(* Logix 5000 project; controller PLC_MCC1300_75F1 vendor 1 type 14 code 166 rev 32.11; software revision 32.04; part 41 of 83 *)
(* tags used below, declared in another part *)
   GP_RampSpace : GP_RampSpace;
   I : INT[128];   // Local Input Updates Input Slot 2
   TMP_d : DINT;
   TMP_dConv : DINT;
   TMP_dConvDebug : DINT;
   TMP_dEndConveyorPos : DINT;
   TMP_dIndexNext : DINT;
   TMP_dIndexNextDebug : DINT;
   TMP_dIndexPreviousDebug : DINT;
   TMP_dTailOnNextConveyor_cmm : DINT;
   TMP_xLastConvDebug : BOOL;
   TMP_xOSN : DINT;
   TMP_xOSN_B : DINT;
   TMP_xOSR : DINT;
   TMP_xOSR_B : DINT;
   xAlwaysOFF : BOOL;
   xAlwaysON : BOOL;
   xDebugOFF : BOOL;
   xDebugON : BOOL;
   Z300_Conveyor : UDT_StandConv[29];
   Z300_Conveyor_ALM : MAC_Conveyor_ZC_ALM[29];
   Z300_Conveyor_Conf : UDT_Conveyor_Config[29];
   Z300_Conveyor_HMR : MAC_Conveyor_ZC_HMR[29];
   Z300_Conveyor_HMW : MAC_Conveyor_ZC_HMW[29];
   Z300_LineTracking : UDT_LINE_TRACKING;
(* MainProgram, continued *)

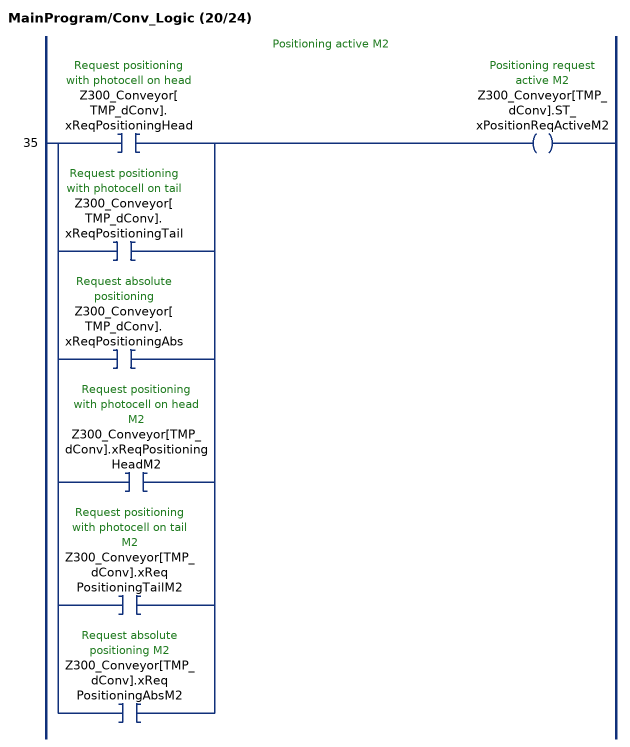
   // Positioning active M2
   35: [XIC(Z300_Conveyor[TMP_dConv].xReqPositioningHead) ,XIC(Z300_Conveyor[TMP_dConv].xReqPositioningTail) ,XIC(Z300_Conveyor[TMP_dConv].xReqPositioningAbs) ,XIC(Z300_Conveyor[TMP_dConv].xReqPositioningHeadM2) ,XIC(Z300_Conveyor[TMP_dConv].xReqPositioningTailM2) ,XIC(Z300_Conveyor[TMP_dConv].xReqPositioningAbsM2) ]OTE(Z300_Conveyor[TMP_dConv].ST_xPositionReqActiveM2);
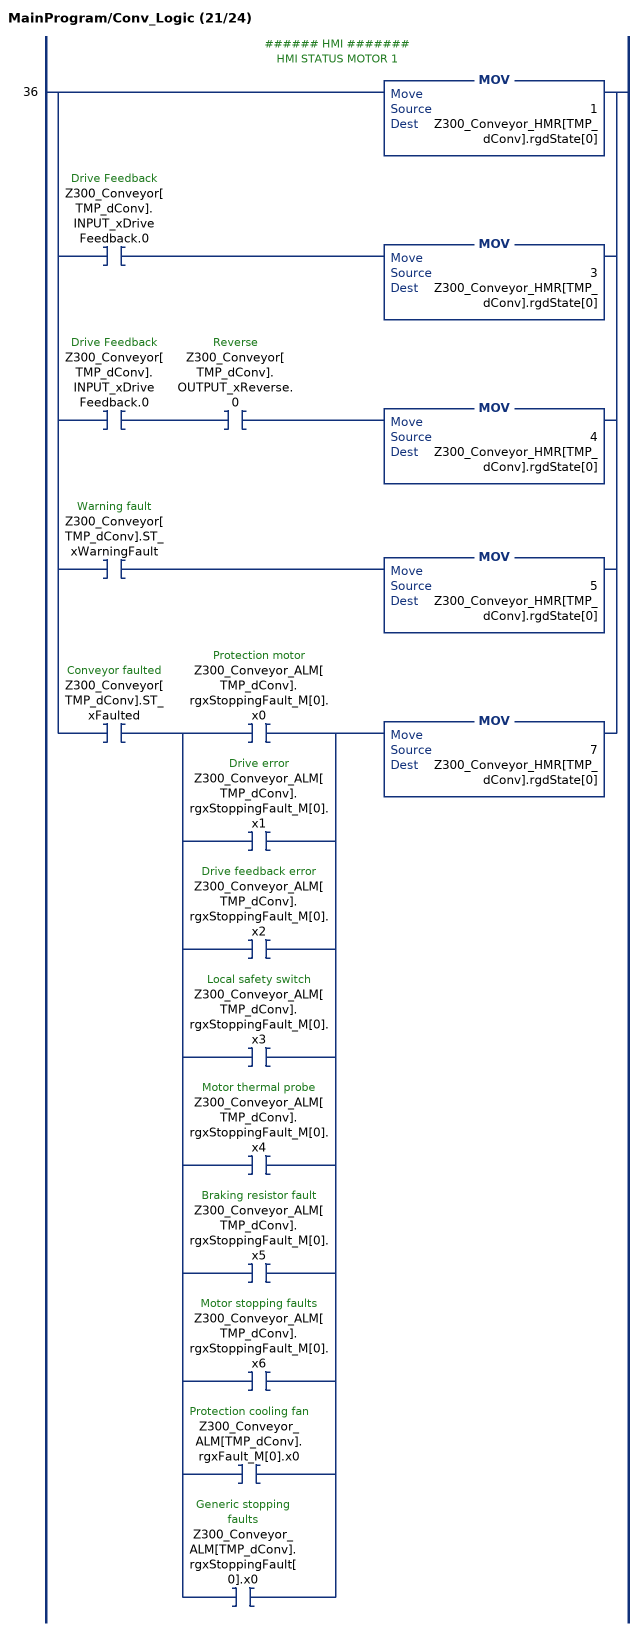
   // ###### HMI #######
   // HMI STATUS MOTOR 1
   36: [MOV(1,Z300_Conveyor_HMR[TMP_dConv].rgdState[0]) ,XIC(Z300_Conveyor[TMP_dConv].INPUT_xDriveFeedback.0) MOV(3,Z300_Conveyor_HMR[TMP_dConv].rgdState[0]) ,XIC(Z300_Conveyor[TMP_dConv].INPUT_xDriveFeedback.0) XIC(Z300_Conveyor[TMP_dConv].OUTPUT_xReverse.0) MOV(4,Z300_Conveyor_HMR[TMP_dConv].rgdState[0]) ,XIC(Z300_Conveyor[TMP_dConv].ST_xWarningFault) MOV(5,Z300_Conveyor_HMR[TMP_dConv].rgdState[0]) ,XIC(Z300_Conveyor[TMP_dConv].ST_xFaulted) [XIC(Z300_Conveyor_ALM[TMP_dConv].rgxStoppingFault_M[0].x0) ,XIC(Z300_Conveyor_ALM[TMP_dConv].rgxStoppingFault_M[0].x1) ,XIC(Z300_Conveyor_ALM[TMP_dConv].rgxStoppingFault_M[0].x2) ,XIC(Z300_Conveyor_ALM[TMP_dConv].rgxStoppingFault_M[0].x3) ,XIC(Z300_Conveyor_ALM[TMP_dConv].rgxStoppingFault_M[0].x4) ,XIC(Z300_Conveyor_ALM[TMP_dConv].rgxStoppingFault_M[0].x5) ,XIC(Z300_Conveyor_ALM[TMP_dConv].rgxStoppingFault_M[0].x6) ,XIC(Z300_Conveyor_ALM[TMP_dConv].rgxFault_M[0].x0) ,XIC(Z300_Conveyor_ALM[TMP_dConv].rgxStoppingFault[0].x0) ] MOV(7,Z300_Conveyor_HMR[TMP_dConv].rgdState[0]) ];
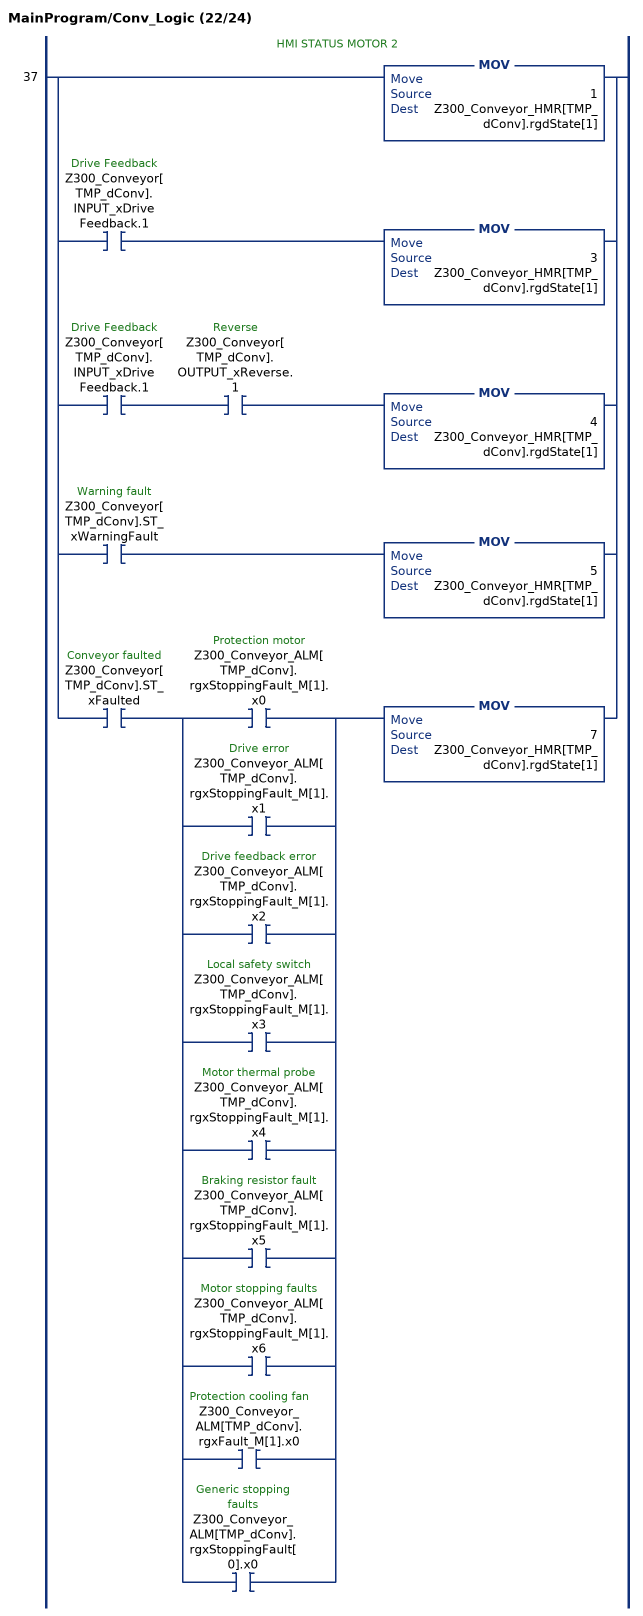
   // HMI STATUS MOTOR 2
   37: [MOV(1,Z300_Conveyor_HMR[TMP_dConv].rgdState[1]) ,XIC(Z300_Conveyor[TMP_dConv].INPUT_xDriveFeedback.1) MOV(3,Z300_Conveyor_HMR[TMP_dConv].rgdState[1]) ,XIC(Z300_Conveyor[TMP_dConv].INPUT_xDriveFeedback.1) XIC(Z300_Conveyor[TMP_dConv].OUTPUT_xReverse.1) MOV(4,Z300_Conveyor_HMR[TMP_dConv].rgdState[1]) ,XIC(Z300_Conveyor[TMP_dConv].ST_xWarningFault) MOV(5,Z300_Conveyor_HMR[TMP_dConv].rgdState[1]) ,XIC(Z300_Conveyor[TMP_dConv].ST_xFaulted) [XIC(Z300_Conveyor_ALM[TMP_dConv].rgxStoppingFault_M[1].x0) ,XIC(Z300_Conveyor_ALM[TMP_dConv].rgxStoppingFault_M[1].x1) ,XIC(Z300_Conveyor_ALM[TMP_dConv].rgxStoppingFault_M[1].x2) ,XIC(Z300_Conveyor_ALM[TMP_dConv].rgxStoppingFault_M[1].x3) ,XIC(Z300_Conveyor_ALM[TMP_dConv].rgxStoppingFault_M[1].x4) ,XIC(Z300_Conveyor_ALM[TMP_dConv].rgxStoppingFault_M[1].x5) ,XIC(Z300_Conveyor_ALM[TMP_dConv].rgxStoppingFault_M[1].x6) ,XIC(Z300_Conveyor_ALM[TMP_dConv].rgxFault_M[1].x0) ,XIC(Z300_Conveyor_ALM[TMP_dConv].rgxStoppingFault[0].x0) ] MOV(7,Z300_Conveyor_HMR[TMP_dConv].rgdState[1]) ];
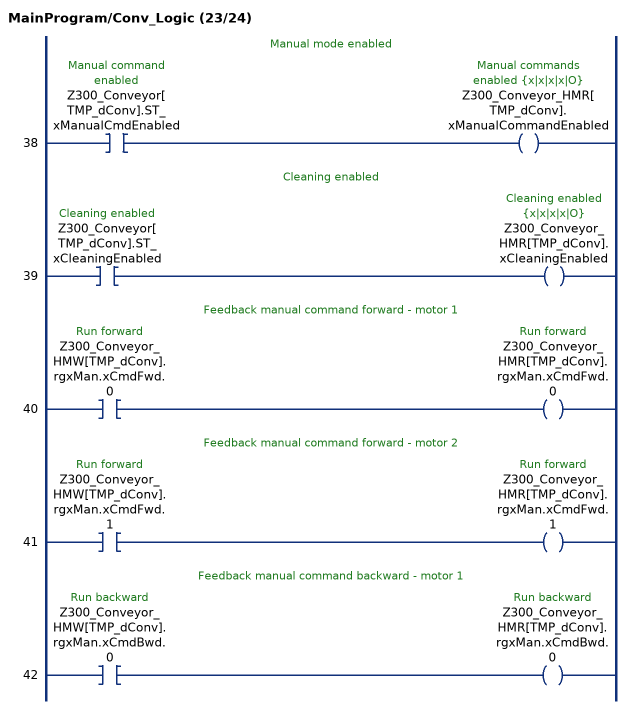
   // Manual mode enabled
   38: XIC(Z300_Conveyor[TMP_dConv].ST_xManualCmdEnabled)OTE(Z300_Conveyor_HMR[TMP_dConv].xManualCommandEnabled);
   // Cleaning enabled
   39: XIC(Z300_Conveyor[TMP_dConv].ST_xCleaningEnabled)OTE(Z300_Conveyor_HMR[TMP_dConv].xCleaningEnabled);
   // Feedback manual command forward - motor 1
   40: XIC(Z300_Conveyor_HMW[TMP_dConv].rgxMan.xCmdFwd.0)OTE(Z300_Conveyor_HMR[TMP_dConv].rgxMan.xCmdFwd.0);
   // Feedback manual command forward - motor 2
   41: XIC(Z300_Conveyor_HMW[TMP_dConv].rgxMan.xCmdFwd.1)OTE(Z300_Conveyor_HMR[TMP_dConv].rgxMan.xCmdFwd.1);
   // Feedback manual command backward - motor 1
   42: XIC(Z300_Conveyor_HMW[TMP_dConv].rgxMan.xCmdBwd.0)OTE(Z300_Conveyor_HMR[TMP_dConv].rgxMan.xCmdBwd.0);
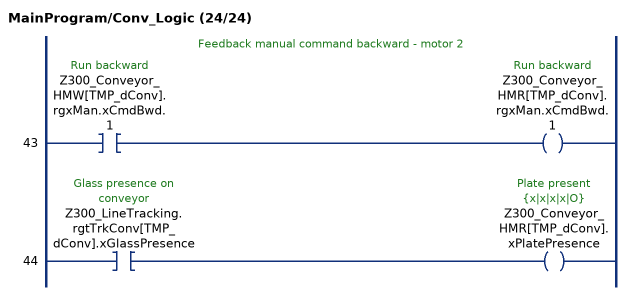
   // Feedback manual command backward - motor 2
   43: XIC(Z300_Conveyor_HMW[TMP_dConv].rgxMan.xCmdBwd.1)OTE(Z300_Conveyor_HMR[TMP_dConv].rgxMan.xCmdBwd.1);
   44: XIC(Z300_LineTracking.rgtTrkConv[TMP_dConv].xGlassPresence)OTE(Z300_Conveyor_HMR[TMP_dConv].xPlatePresence);
END_ROUTINE

ROUTINE Conv_Logic_Debug   (* ladder *)
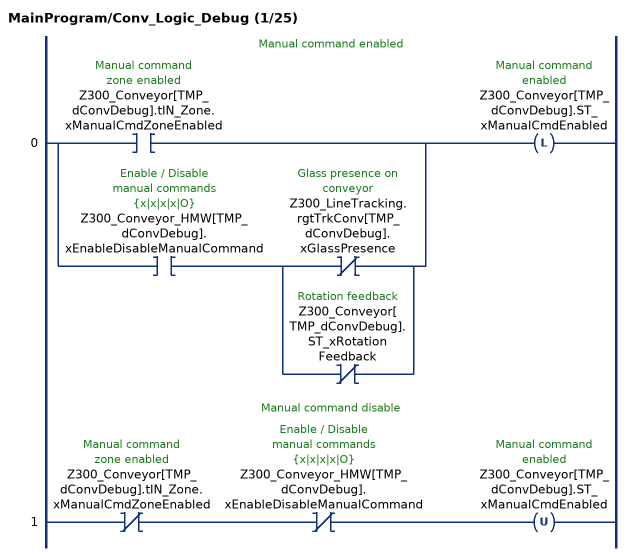
   // Manual command enabled
   0: [XIC(Z300_Conveyor[TMP_dConvDebug].tIN_Zone.xManualCmdZoneEnabled) ,XIC(Z300_Conveyor_HMW[TMP_dConvDebug].xEnableDisableManualCommand) [XIO(Z300_LineTracking.rgtTrkConv[TMP_dConvDebug].xGlassPresence) ,XIO(Z300_Conveyor[TMP_dConvDebug].ST_xRotationFeedback) ] ]OTL(Z300_Conveyor[TMP_dConvDebug].ST_xManualCmdEnabled);
   // Manual command disable
   1: XIO(Z300_Conveyor[TMP_dConvDebug].tIN_Zone.xManualCmdZoneEnabled)XIO(Z300_Conveyor_HMW[TMP_dConvDebug].xEnableDisableManualCommand)OTU(Z300_Conveyor[TMP_dConvDebug].ST_xManualCmdEnabled);
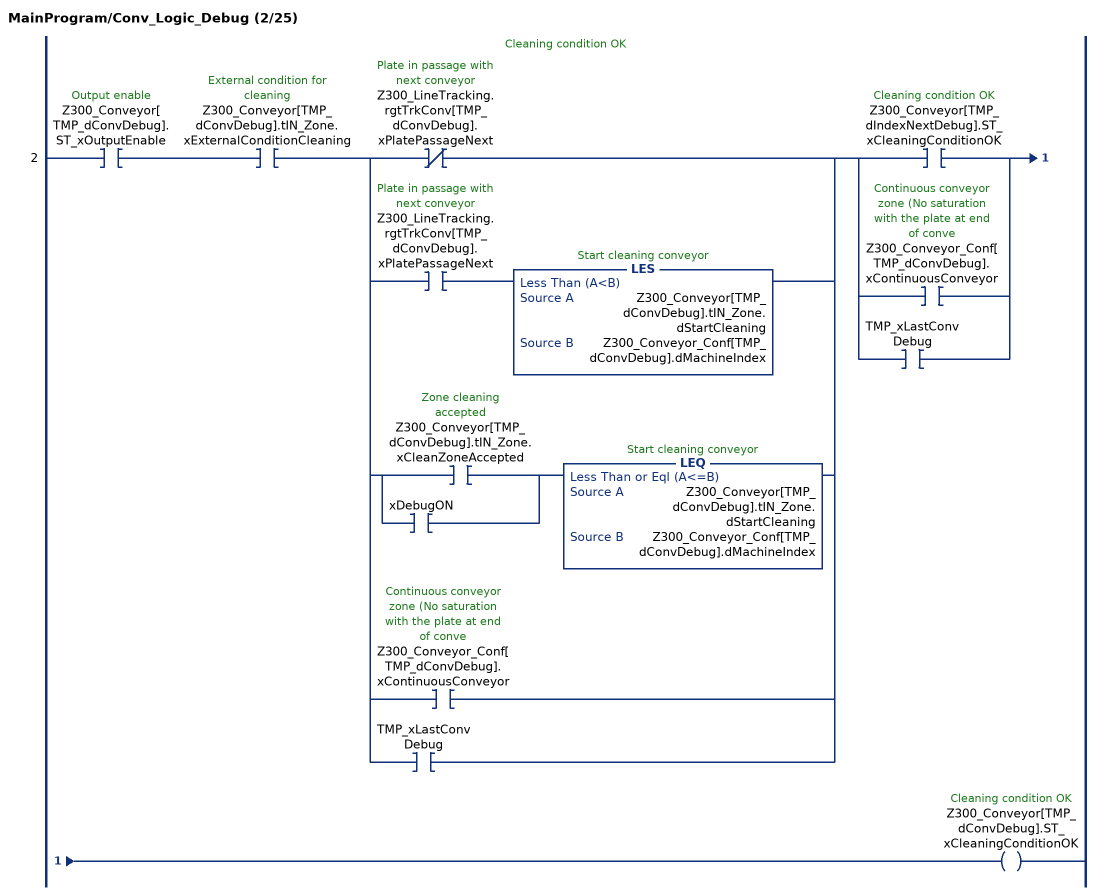
   // Cleaning condition OK
   2: XIC(Z300_Conveyor[TMP_dConvDebug].ST_xOutputEnable)XIC(Z300_Conveyor[TMP_dConvDebug].tIN_Zone.xExternalConditionCleaning)[[XIO(Z300_LineTracking.rgtTrkConv[TMP_dConvDebug].xPlatePassageNext) ,XIC(Z300_LineTracking.rgtTrkConv[TMP_dConvDebug].xPlatePassageNext) LES(Z300_Conveyor[TMP_dConvDebug].tIN_Zone.dStartCleaning,Z300_Conveyor_Conf[TMP_dConvDebug].dMachineIndex) ] ,[[XIC(Z300_Conveyor[TMP_dConvDebug].tIN_Zone.xCleanZoneAccepted) ,XIC(xDebugON) ] LEQ(Z300_Conveyor[TMP_dConvDebug].tIN_Zone.dStartCleaning,Z300_Conveyor_Conf[TMP_dConvDebug].dMachineIndex) ,XIC(Z300_Conveyor_Conf[TMP_dConvDebug].xContinuousConveyor) ,XIC(TMP_xLastConvDebug) ] ][XIC(Z300_Conveyor[TMP_dIndexNextDebug].ST_xCleaningConditionOK) ,XIC(Z300_Conveyor_Conf[TMP_dConvDebug].xContinuousConveyor) ,XIC(TMP_xLastConvDebug) ]OTE(Z300_Conveyor[TMP_dConvDebug].ST_xCleaningConditionOK);
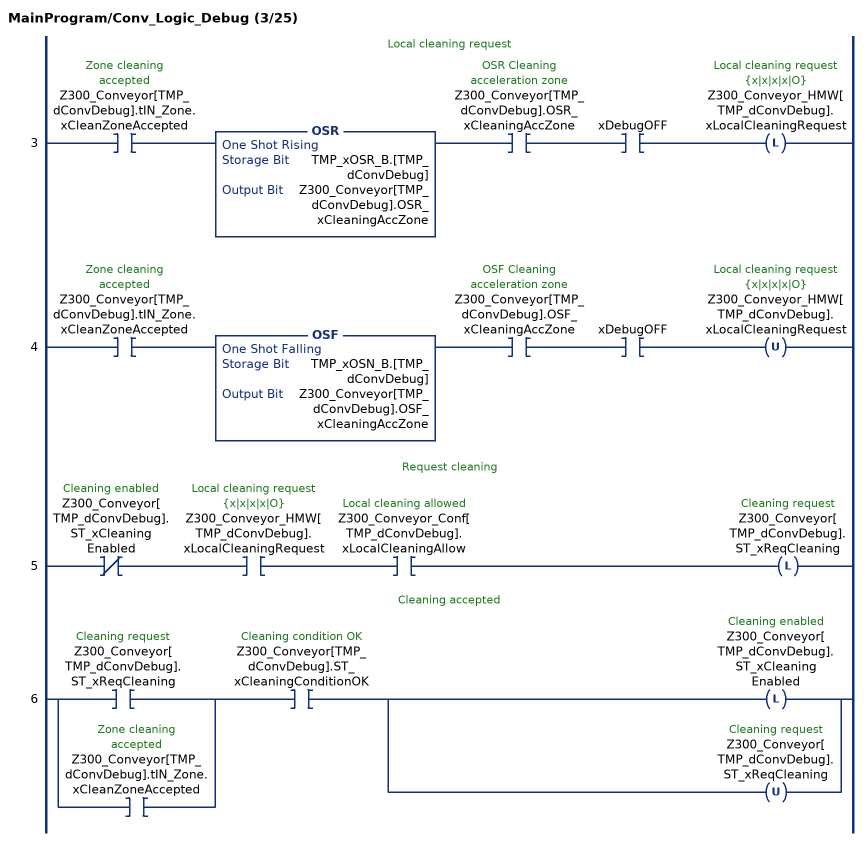
   // Local cleaning request
   3: XIC(Z300_Conveyor[TMP_dConvDebug].tIN_Zone.xCleanZoneAccepted)OSR(TMP_xOSR_B.[TMP_dConvDebug],Z300_Conveyor[TMP_dConvDebug].OSR_xCleaningAccZone)XIC(Z300_Conveyor[TMP_dConvDebug].OSR_xCleaningAccZone)XIC(xDebugOFF)OTL(Z300_Conveyor_HMW[TMP_dConvDebug].xLocalCleaningRequest);
   4: XIC(Z300_Conveyor[TMP_dConvDebug].tIN_Zone.xCleanZoneAccepted)OSF(TMP_xOSN_B.[TMP_dConvDebug],Z300_Conveyor[TMP_dConvDebug].OSF_xCleaningAccZone)XIC(Z300_Conveyor[TMP_dConvDebug].OSF_xCleaningAccZone)XIC(xDebugOFF)OTU(Z300_Conveyor_HMW[TMP_dConvDebug].xLocalCleaningRequest);
   // Request cleaning
   5: XIO(Z300_Conveyor[TMP_dConvDebug].ST_xCleaningEnabled)XIC(Z300_Conveyor_HMW[TMP_dConvDebug].xLocalCleaningRequest)XIC(Z300_Conveyor_Conf[TMP_dConvDebug].xLocalCleaningAllow)OTL(Z300_Conveyor[TMP_dConvDebug].ST_xReqCleaning);
   // Cleaning accepted
   6: [XIC(Z300_Conveyor[TMP_dConvDebug].ST_xReqCleaning) ,XIC(Z300_Conveyor[TMP_dConvDebug].tIN_Zone.xCleanZoneAccepted) ]XIC(Z300_Conveyor[TMP_dConvDebug].ST_xCleaningConditionOK)[OTL(Z300_Conveyor[TMP_dConvDebug].ST_xCleaningEnabled) ,OTU(Z300_Conveyor[TMP_dConvDebug].ST_xReqCleaning) ];
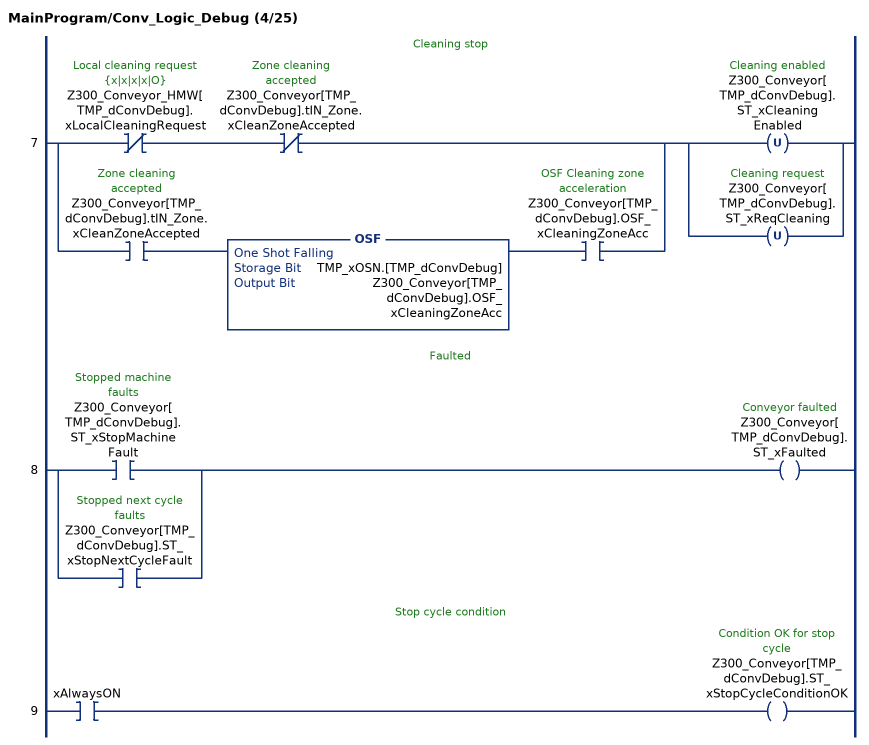
   // Cleaning stop
   7: [XIO(Z300_Conveyor_HMW[TMP_dConvDebug].xLocalCleaningRequest) XIO(Z300_Conveyor[TMP_dConvDebug].tIN_Zone.xCleanZoneAccepted) ,XIC(Z300_Conveyor[TMP_dConvDebug].tIN_Zone.xCleanZoneAccepted) OSF(TMP_xOSN.[TMP_dConvDebug],Z300_Conveyor[TMP_dConvDebug].OSF_xCleaningZoneAcc) XIC(Z300_Conveyor[TMP_dConvDebug].OSF_xCleaningZoneAcc) ][OTU(Z300_Conveyor[TMP_dConvDebug].ST_xCleaningEnabled) ,OTU(Z300_Conveyor[TMP_dConvDebug].ST_xReqCleaning) ];
   // Faulted
   8: [XIC(Z300_Conveyor[TMP_dConvDebug].ST_xStopMachineFault) ,XIC(Z300_Conveyor[TMP_dConvDebug].ST_xStopNextCycleFault) ]OTE(Z300_Conveyor[TMP_dConvDebug].ST_xFaulted);
   // Stop cycle condition
   9: XIC(xAlwaysON)OTE(Z300_Conveyor[TMP_dConvDebug].ST_xStopCycleConditionOK);
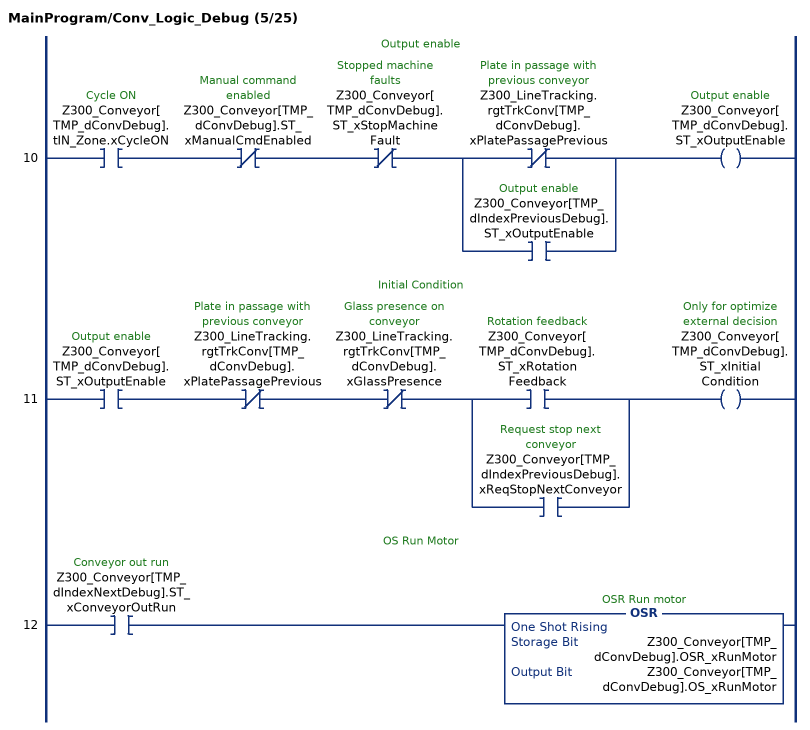
   // Output enable
   10: XIC(Z300_Conveyor[TMP_dConvDebug].tIN_Zone.xCycleON)XIO(Z300_Conveyor[TMP_dConvDebug].ST_xManualCmdEnabled)XIO(Z300_Conveyor[TMP_dConvDebug].ST_xStopMachineFault)[XIO(Z300_LineTracking.rgtTrkConv[TMP_dConvDebug].xPlatePassagePrevious) ,XIC(Z300_Conveyor[TMP_dIndexPreviousDebug].ST_xOutputEnable) ]OTE(Z300_Conveyor[TMP_dConvDebug].ST_xOutputEnable);
   // Initial Condition
   11: XIC(Z300_Conveyor[TMP_dConvDebug].ST_xOutputEnable)XIO(Z300_LineTracking.rgtTrkConv[TMP_dConvDebug].xPlatePassagePrevious)XIO(Z300_LineTracking.rgtTrkConv[TMP_dConvDebug].xGlassPresence)[XIC(Z300_Conveyor[TMP_dConvDebug].ST_xRotationFeedback) ,XIC(Z300_Conveyor[TMP_dIndexPreviousDebug].xReqStopNextConveyor) ]OTE(Z300_Conveyor[TMP_dConvDebug].ST_xInitialCondition);
   // OS Run Motor
   12: XIC(Z300_Conveyor[TMP_dIndexNextDebug].ST_xConveyorOutRun)OSR(Z300_Conveyor[TMP_dConvDebug].OSR_xRunMotor,Z300_Conveyor[TMP_dConvDebug].OS_xRunMotor);
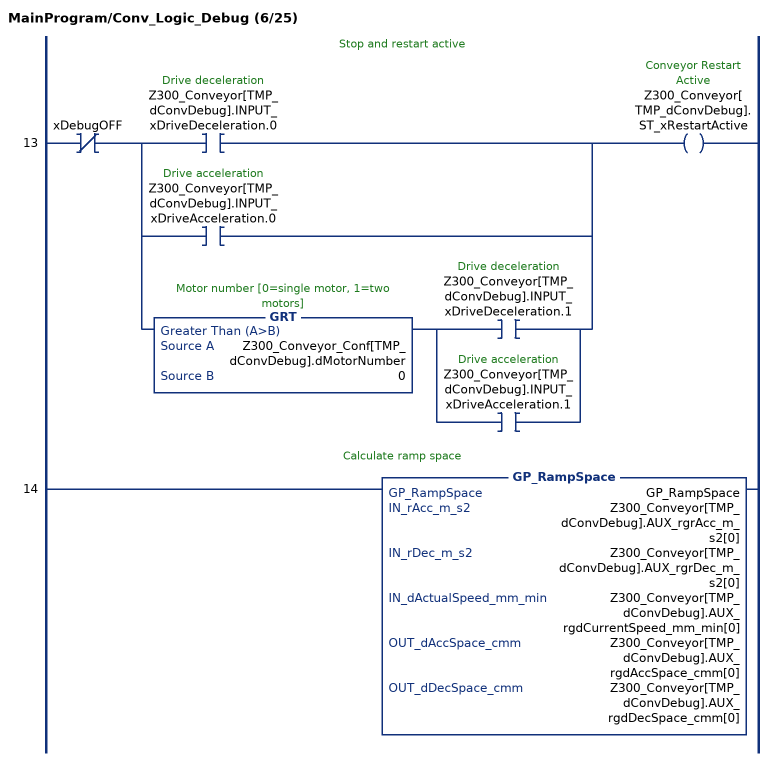
   // Stop and restart active
   13: XIO(xDebugOFF)[[XIC(Z300_Conveyor[TMP_dConvDebug].INPUT_xDriveDeceleration.0) ,XIC(Z300_Conveyor[TMP_dConvDebug].INPUT_xDriveAcceleration.0) ] ,GRT(Z300_Conveyor_Conf[TMP_dConvDebug].dMotorNumber,0) [XIC(Z300_Conveyor[TMP_dConvDebug].INPUT_xDriveDeceleration.1) ,XIC(Z300_Conveyor[TMP_dConvDebug].INPUT_xDriveAcceleration.1) ] ]OTE(Z300_Conveyor[TMP_dConvDebug].ST_xRestartActive);
   // Calculate ramp space
   14: GP_RampSpace(GP_RampSpace,Z300_Conveyor[TMP_dConvDebug].AUX_rgrAcc_m_s2[0],Z300_Conveyor[TMP_dConvDebug].AUX_rgrDec_m_s2[0],Z300_Conveyor[TMP_dConvDebug].AUX_rgdCurrentSpeed_mm_min[0],Z300_Conveyor[TMP_dConvDebug].AUX_rgdAccSpace_cmm[0],Z300_Conveyor[TMP_dConvDebug].AUX_rgdDecSpace_cmm[0]);
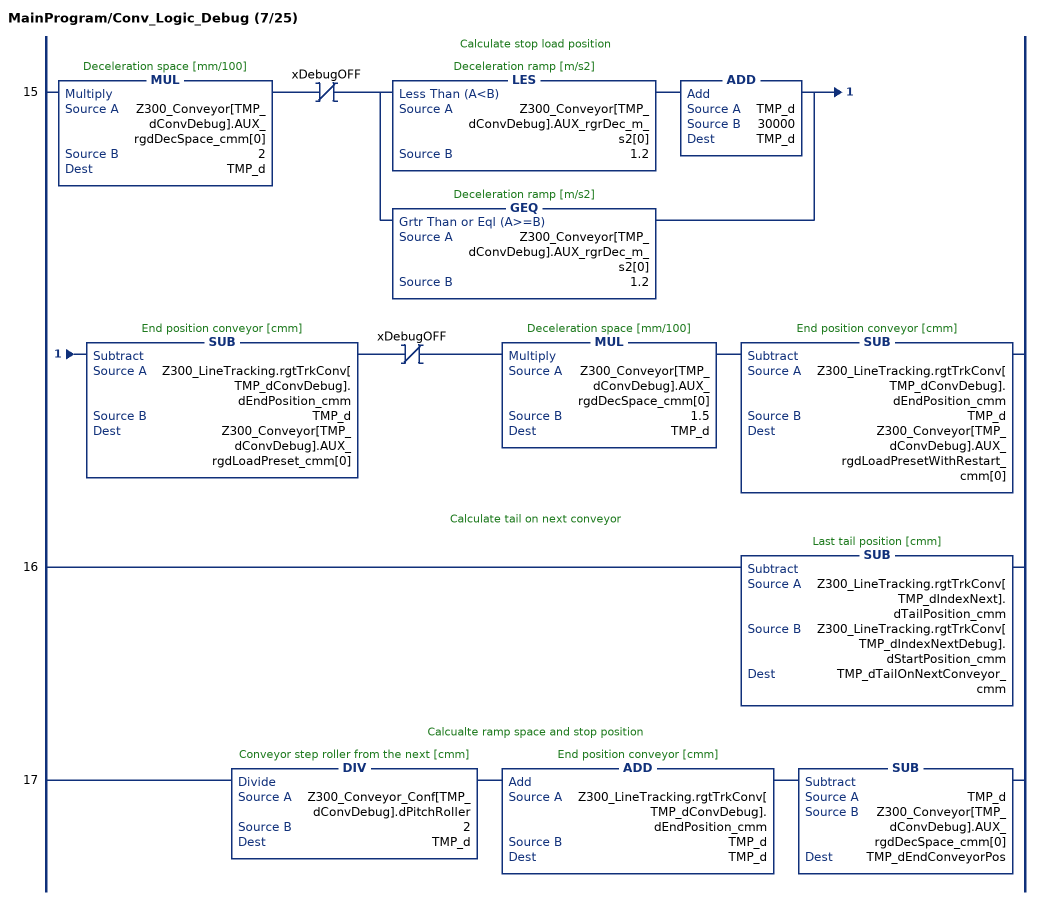
   // Calculate stop load position
   15: MUL(Z300_Conveyor[TMP_dConvDebug].AUX_rgdDecSpace_cmm[0],2,TMP_d)XIO(xDebugOFF)[LES(Z300_Conveyor[TMP_dConvDebug].AUX_rgrDec_m_s2[0],1.2) ADD(TMP_d,30000,TMP_d) ,GEQ(Z300_Conveyor[TMP_dConvDebug].AUX_rgrDec_m_s2[0],1.2) ]SUB(Z300_LineTracking.rgtTrkConv[TMP_dConvDebug].dEndPosition_cmm,TMP_d,Z300_Conveyor[TMP_dConvDebug].AUX_rgdLoadPreset_cmm[0])XIO(xDebugOFF)MUL(Z300_Conveyor[TMP_dConvDebug].AUX_rgdDecSpace_cmm[0],1.5,TMP_d)SUB(Z300_LineTracking.rgtTrkConv[TMP_dConvDebug].dEndPosition_cmm,TMP_d,Z300_Conveyor[TMP_dConvDebug].AUX_rgdLoadPresetWithRestart_cmm[0]);
   // Calculate tail on next conveyor
   16: SUB(Z300_LineTracking.rgtTrkConv[TMP_dIndexNext].dTailPosition_cmm,Z300_LineTracking.rgtTrkConv[TMP_dIndexNextDebug].dStartPosition_cmm,TMP_dTailOnNextConveyor_cmm);
   // Calcualte ramp space and stop position
   17: DIV(Z300_Conveyor_Conf[TMP_dConvDebug].dPitchRoller,2,TMP_d)ADD(Z300_LineTracking.rgtTrkConv[TMP_dConvDebug].dEndPosition_cmm,TMP_d,TMP_d)SUB(TMP_d,Z300_Conveyor[TMP_dConvDebug].AUX_rgdDecSpace_cmm[0],TMP_dEndConveyorPos);
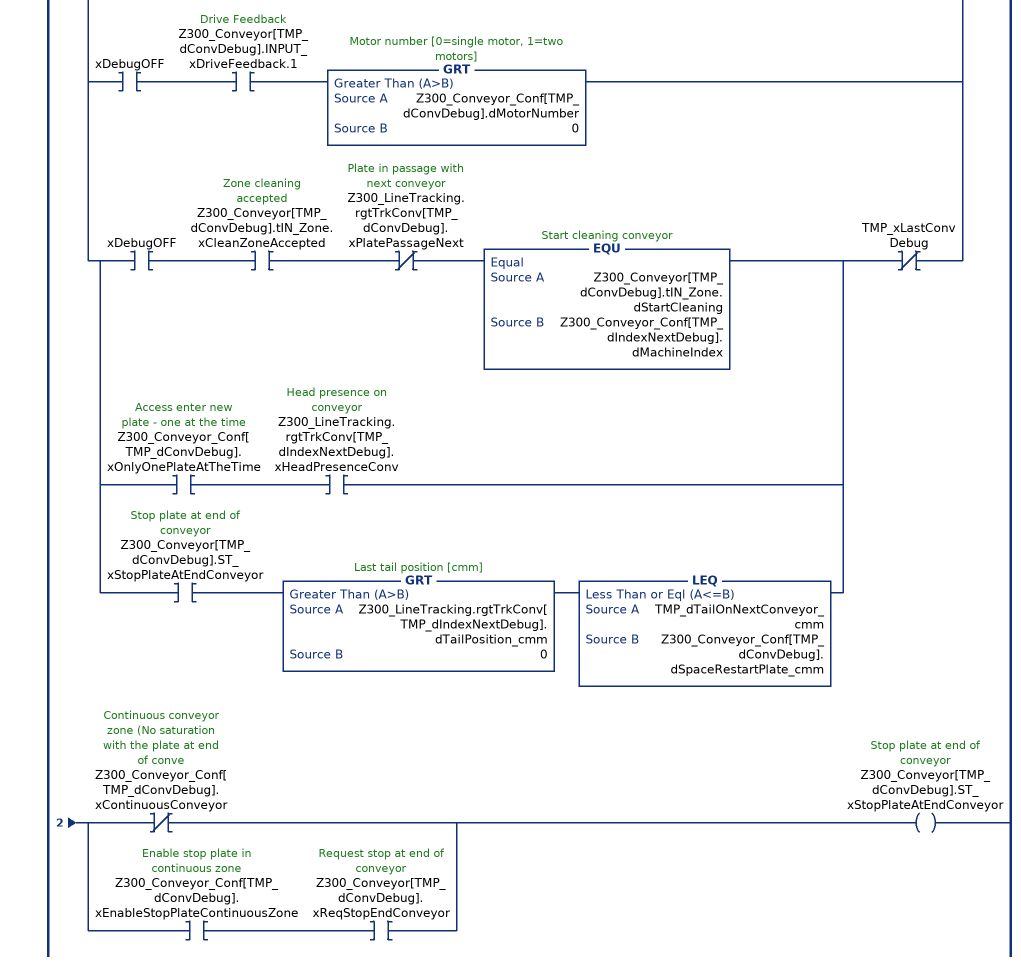
   // Stop at end of conveyor if next not run
   18: [GEQ(Z300_LineTracking.rgtTrkConv[TMP_dConvDebug].dHeadPosition_cmm,Z300_Conveyor[TMP_dConvDebug].AUX_rgdLoadPreset_cmm[0]) ,XIC(Z300_Conveyor[TMP_dConvDebug].ST_xStopPlateAtEndConveyor) XIC(Z300_LineTracking.rgtTrkConv[TMP_dConvDebug].xGlassPresCom) ][[XIO(Z300_Conveyor[TMP_dIndexNextDebug].ST_xConveyorOutRun) ,XIC(xDebugON) ] [XIO(Z300_Conveyor[TMP_dIndexNextDebug].ST_rgxConveyorOutRunSgm.0) ,XIO(Z300_Conveyor[TMP_dIndexNextDebug].ST_rgxConveyorOutRunSgm.1) GRT(Z300_Conveyor_Conf[TMP_dIndexNextDebug].dMotorNumber,0) ] XIO(TMP_xLastConvDebug) ,XIC(Z300_Conveyor[TMP_dIndexNextDebug].xReqExtStopLoadNewPlate) ,XIO(Z300_Conveyor[TMP_dConvDebug].ST_xCleaningEnabled) XIC(Z300_Conveyor[TMP_dIndexNextDebug].ST_xCleaningEnabled) XIO(Z300_LineTracking.rgtTrkConv[TMP_dConvDebug].xPlatePassageNext) ,XIC(Z300_Conveyor[TMP_dConvDebug].xReqStopEndConveyor) ,XIC(xDebugOFF) XIC(Z300_Conveyor[TMP_dConvDebug].INPUT_xDriveFeedback.0) ,XIC(xDebugOFF) XIC(Z300_Conveyor[TMP_dConvDebug].INPUT_xDriveFeedback.1) GRT(Z300_Conveyor_Conf[TMP_dConvDebug].dMotorNumber,0) ,[XIC(xDebugOFF) XIC(Z300_Conveyor[TMP_dConvDebug].tIN_Zone.xCleanZoneAccepted) XIO(Z300_LineTracking.rgtTrkConv[TMP_dConvDebug].xPlatePassageNext) EQU(Z300_Conveyor[TMP_dConvDebug].tIN_Zone.dStartCleaning,Z300_Conveyor_Conf[TMP_dIndexNextDebug].dMachineIndex) ,XIC(Z300_Conveyor_Conf[TMP_dConvDebug].xOnlyOnePlateAtTheTime) XIC(Z300_LineTracking.rgtTrkConv[TMP_dIndexNextDebug].xHeadPresenceConv) ,XIC(Z300_Conveyor[TMP_dConvDebug].ST_xStopPlateAtEndConveyor) GRT(Z300_LineTracking.rgtTrkConv[TMP_dIndexNextDebug].dTailPosition_cmm,0) LEQ(TMP_dTailOnNextConveyor_cmm,Z300_Conveyor_Conf[TMP_dConvDebug].dSpaceRestartPlate_cmm) ] XIO(TMP_xLastConvDebug) ][XIO(Z300_Conveyor_Conf[TMP_dConvDebug].xContinuousConveyor) ,XIC(Z300_Conveyor_Conf[TMP_dConvDebug].xEnableStopPlateContinuousZone) XIC(Z300_Conveyor[TMP_dConvDebug].xReqStopEndConveyor) ]OTE(Z300_Conveyor[TMP_dConvDebug].ST_xStopPlateAtEndConveyor);